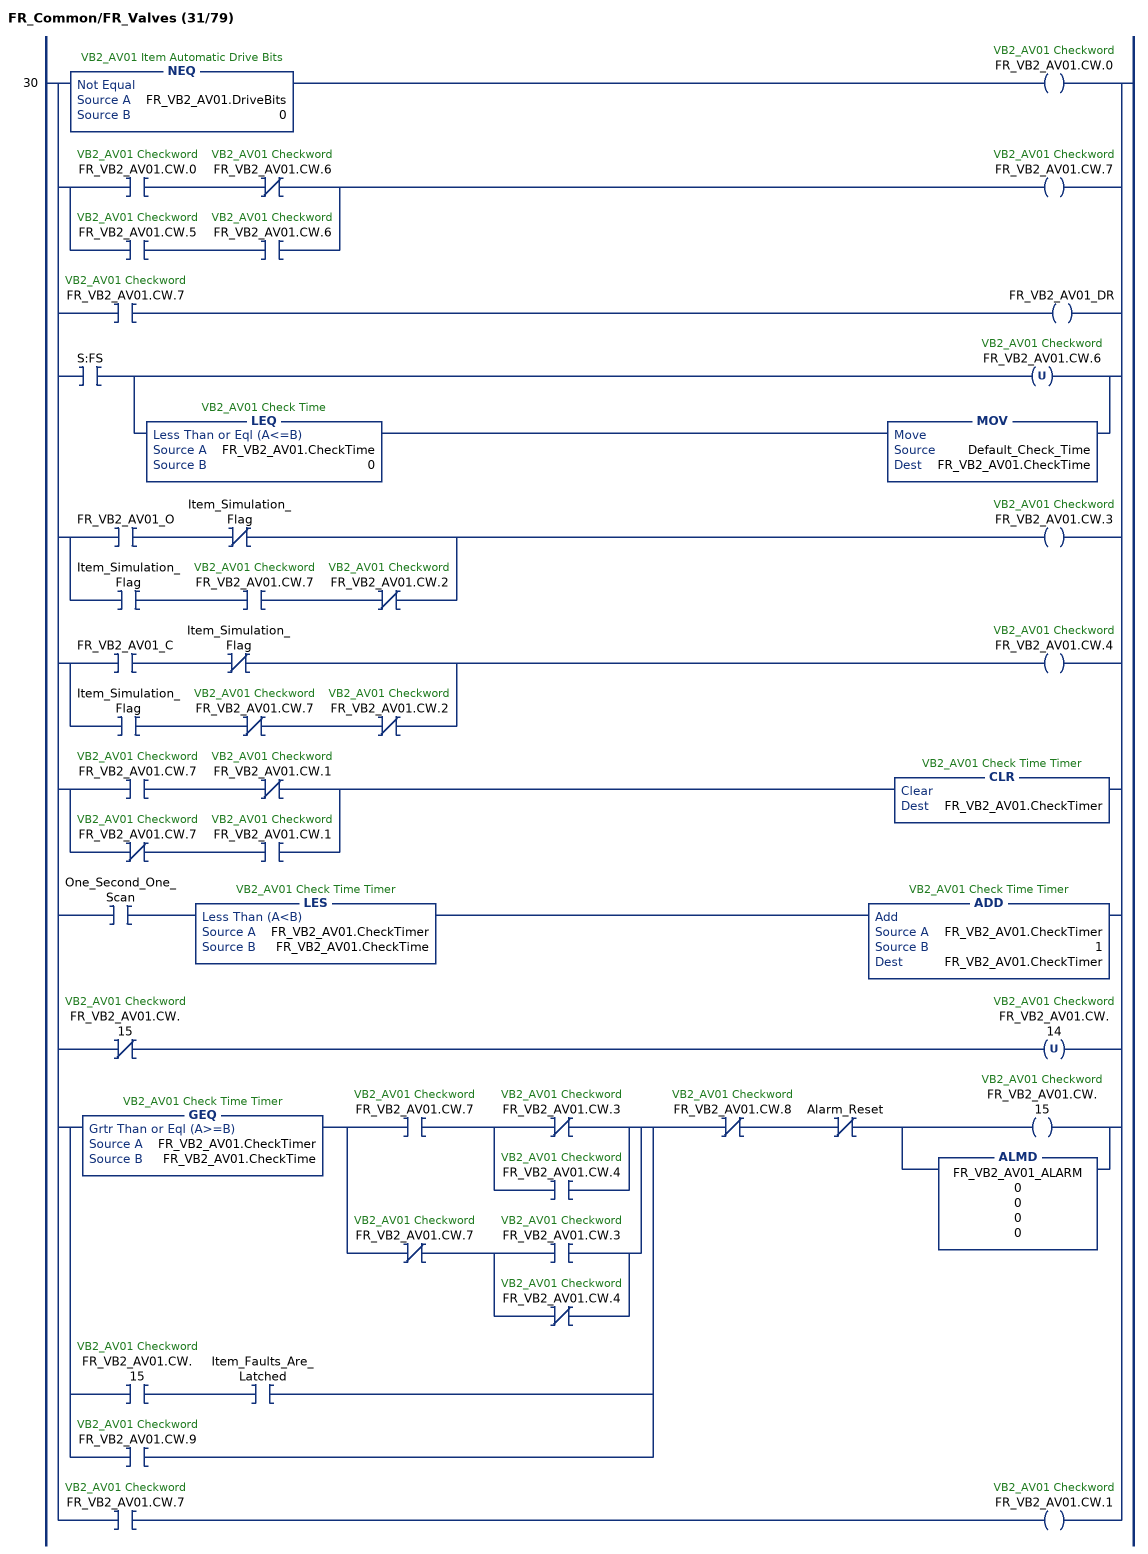
   30: [NEQ(FR_VB2_AV01.DriveBits,0) OTE(FR_VB2_AV01.CW.0) ,[XIC(FR_VB2_AV01.CW.0) XIO(FR_VB2_AV01.CW.6) ,XIC(FR_VB2_AV01.CW.5) XIC(FR_VB2_AV01.CW.6) ] OTE(FR_VB2_AV01.CW.7) ,XIC(FR_VB2_AV01.CW.7) OTE(FR_VB2_AV01_DR) ,XIC(S:FS) [OTU(FR_VB2_AV01.CW.6) ,LEQ(FR_VB2_AV01.CheckTime,0) MOV(Default_Check_Time,FR_VB2_AV01.CheckTime) ] ,[[XIC(FR_VB2_AV01_O) XIO(Item_Simulation_Flag) ,XIC(Item_Simulation_Flag) XIC(FR_VB2_AV01.CW.7) XIO(FR_VB2_AV01.CW.2) ] OTE(FR_VB2_AV01.CW.3) ,[XIC(FR_VB2_AV01_C) XIO(Item_Simulation_Flag) ,XIC(Item_Simulation_Flag) XIO(FR_VB2_AV01.CW.7) XIO(FR_VB2_AV01.CW.2) ] OTE(FR_VB2_AV01.CW.4) ] ,[XIC(FR_VB2_AV01.CW.7) XIO(FR_VB2_AV01.CW.1) ,XIO(FR_VB2_AV01.CW.7) XIC(FR_VB2_AV01.CW.1) ] CLR(FR_VB2_AV01.CheckTimer) ,XIC(One_Second_One_Scan) LES(FR_VB2_AV01.CheckTimer,FR_VB2_AV01.CheckTime) ADD(FR_VB2_AV01.CheckTimer,1,FR_VB2_AV01.CheckTimer) ,XIO(FR_VB2_AV01.CW.15) OTU(FR_VB2_AV01.CW.14) ,[GEQ(FR_VB2_AV01.CheckTimer,FR_VB2_AV01.CheckTime) [XIC(FR_VB2_AV01.CW.7) [XIO(FR_VB2_AV01.CW.3) ,XIC(FR_VB2_AV01.CW.4) ] ,XIO(FR_VB2_AV01.CW.7) [XIC(FR_VB2_AV01.CW.3) ,XIO(FR_VB2_AV01.CW.4) ] ] ,XIC(FR_VB2_AV01.CW.15) XIC(Item_Faults_Are_Latched) ,XIC(FR_VB2_AV01.CW.9) ] XIO(FR_VB2_AV01.CW.8) XIO(Alarm_Reset) [OTE(FR_VB2_AV01.CW.15) ,ALMD(FR_VB2_AV01_ALARM,0,0,0,0) ] ,XIC(FR_VB2_AV01.CW.7) OTE(FR_VB2_AV01.CW.1) ];
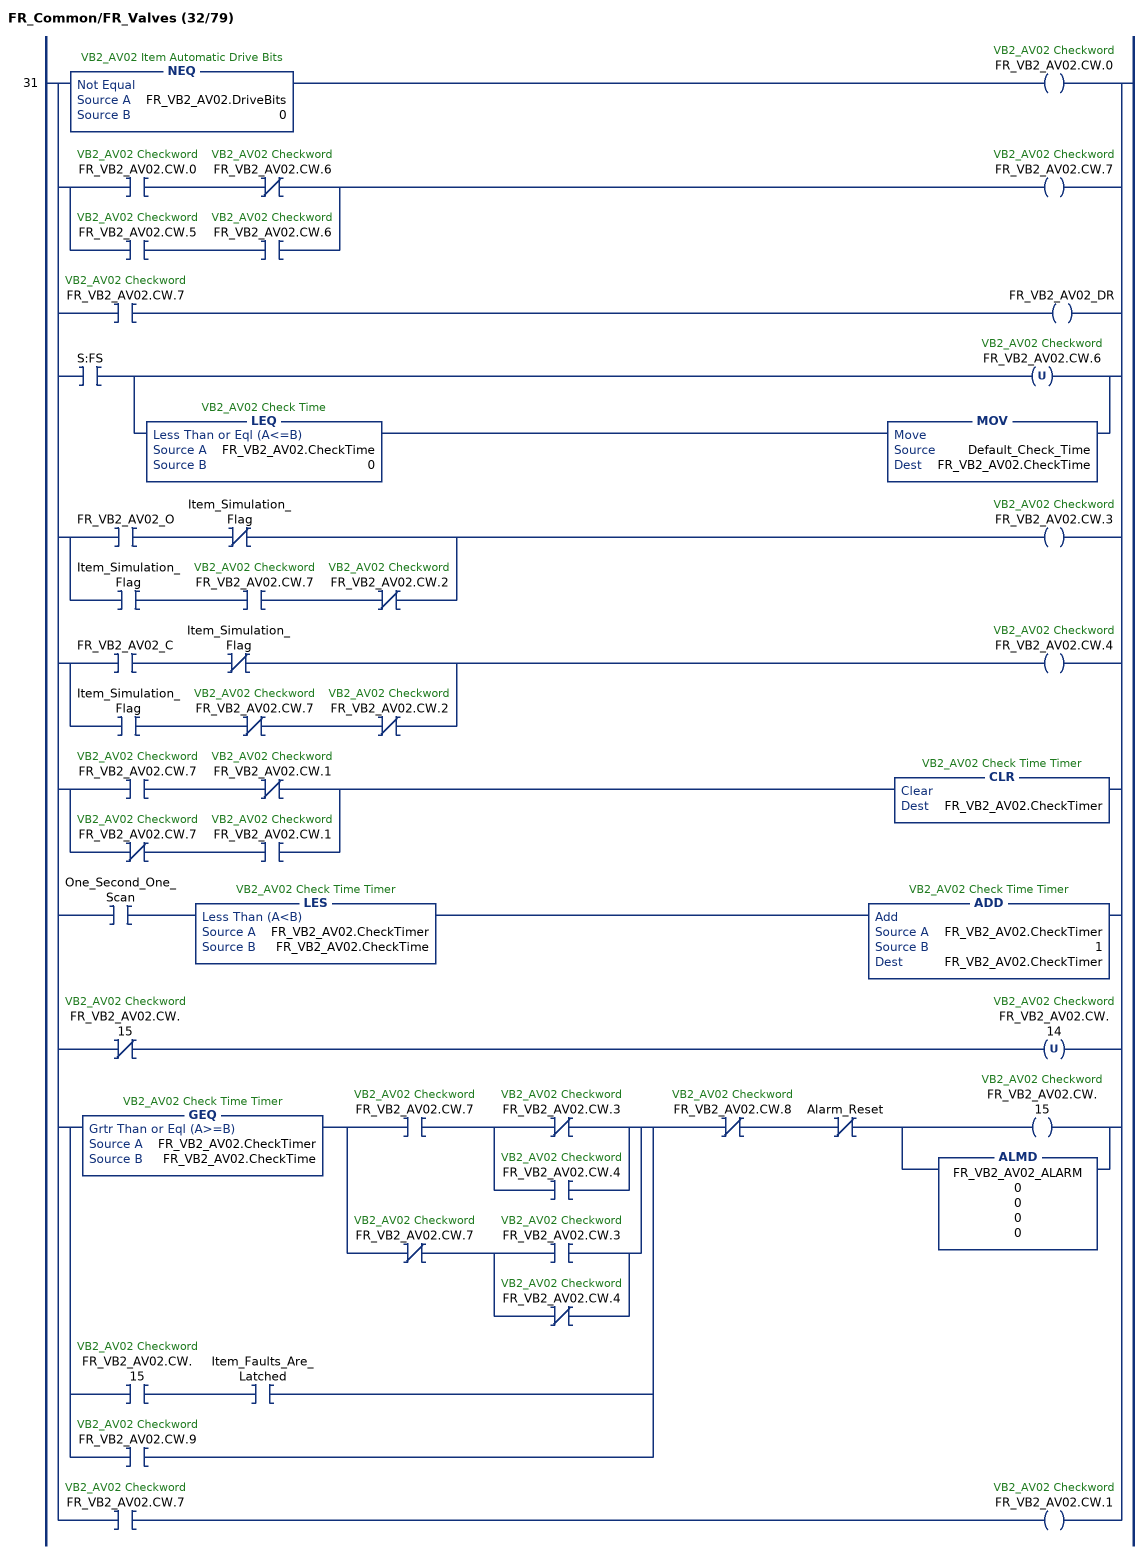
   31: [NEQ(FR_VB2_AV02.DriveBits,0) OTE(FR_VB2_AV02.CW.0) ,[XIC(FR_VB2_AV02.CW.0) XIO(FR_VB2_AV02.CW.6) ,XIC(FR_VB2_AV02.CW.5) XIC(FR_VB2_AV02.CW.6) ] OTE(FR_VB2_AV02.CW.7) ,XIC(FR_VB2_AV02.CW.7) OTE(FR_VB2_AV02_DR) ,XIC(S:FS) [OTU(FR_VB2_AV02.CW.6) ,LEQ(FR_VB2_AV02.CheckTime,0) MOV(Default_Check_Time,FR_VB2_AV02.CheckTime) ] ,[[XIC(FR_VB2_AV02_O) XIO(Item_Simulation_Flag) ,XIC(Item_Simulation_Flag) XIC(FR_VB2_AV02.CW.7) XIO(FR_VB2_AV02.CW.2) ] OTE(FR_VB2_AV02.CW.3) ,[XIC(FR_VB2_AV02_C) XIO(Item_Simulation_Flag) ,XIC(Item_Simulation_Flag) XIO(FR_VB2_AV02.CW.7) XIO(FR_VB2_AV02.CW.2) ] OTE(FR_VB2_AV02.CW.4) ] ,[XIC(FR_VB2_AV02.CW.7) XIO(FR_VB2_AV02.CW.1) ,XIO(FR_VB2_AV02.CW.7) XIC(FR_VB2_AV02.CW.1) ] CLR(FR_VB2_AV02.CheckTimer) ,XIC(One_Second_One_Scan) LES(FR_VB2_AV02.CheckTimer,FR_VB2_AV02.CheckTime) ADD(FR_VB2_AV02.CheckTimer,1,FR_VB2_AV02.CheckTimer) ,XIO(FR_VB2_AV02.CW.15) OTU(FR_VB2_AV02.CW.14) ,[GEQ(FR_VB2_AV02.CheckTimer,FR_VB2_AV02.CheckTime) [XIC(FR_VB2_AV02.CW.7) [XIO(FR_VB2_AV02.CW.3) ,XIC(FR_VB2_AV02.CW.4) ] ,XIO(FR_VB2_AV02.CW.7) [XIC(FR_VB2_AV02.CW.3) ,XIO(FR_VB2_AV02.CW.4) ] ] ,XIC(FR_VB2_AV02.CW.15) XIC(Item_Faults_Are_Latched) ,XIC(FR_VB2_AV02.CW.9) ] XIO(FR_VB2_AV02.CW.8) XIO(Alarm_Reset) [OTE(FR_VB2_AV02.CW.15) ,ALMD(FR_VB2_AV02_ALARM,0,0,0,0) ] ,XIC(FR_VB2_AV02.CW.7) OTE(FR_VB2_AV02.CW.1) ];
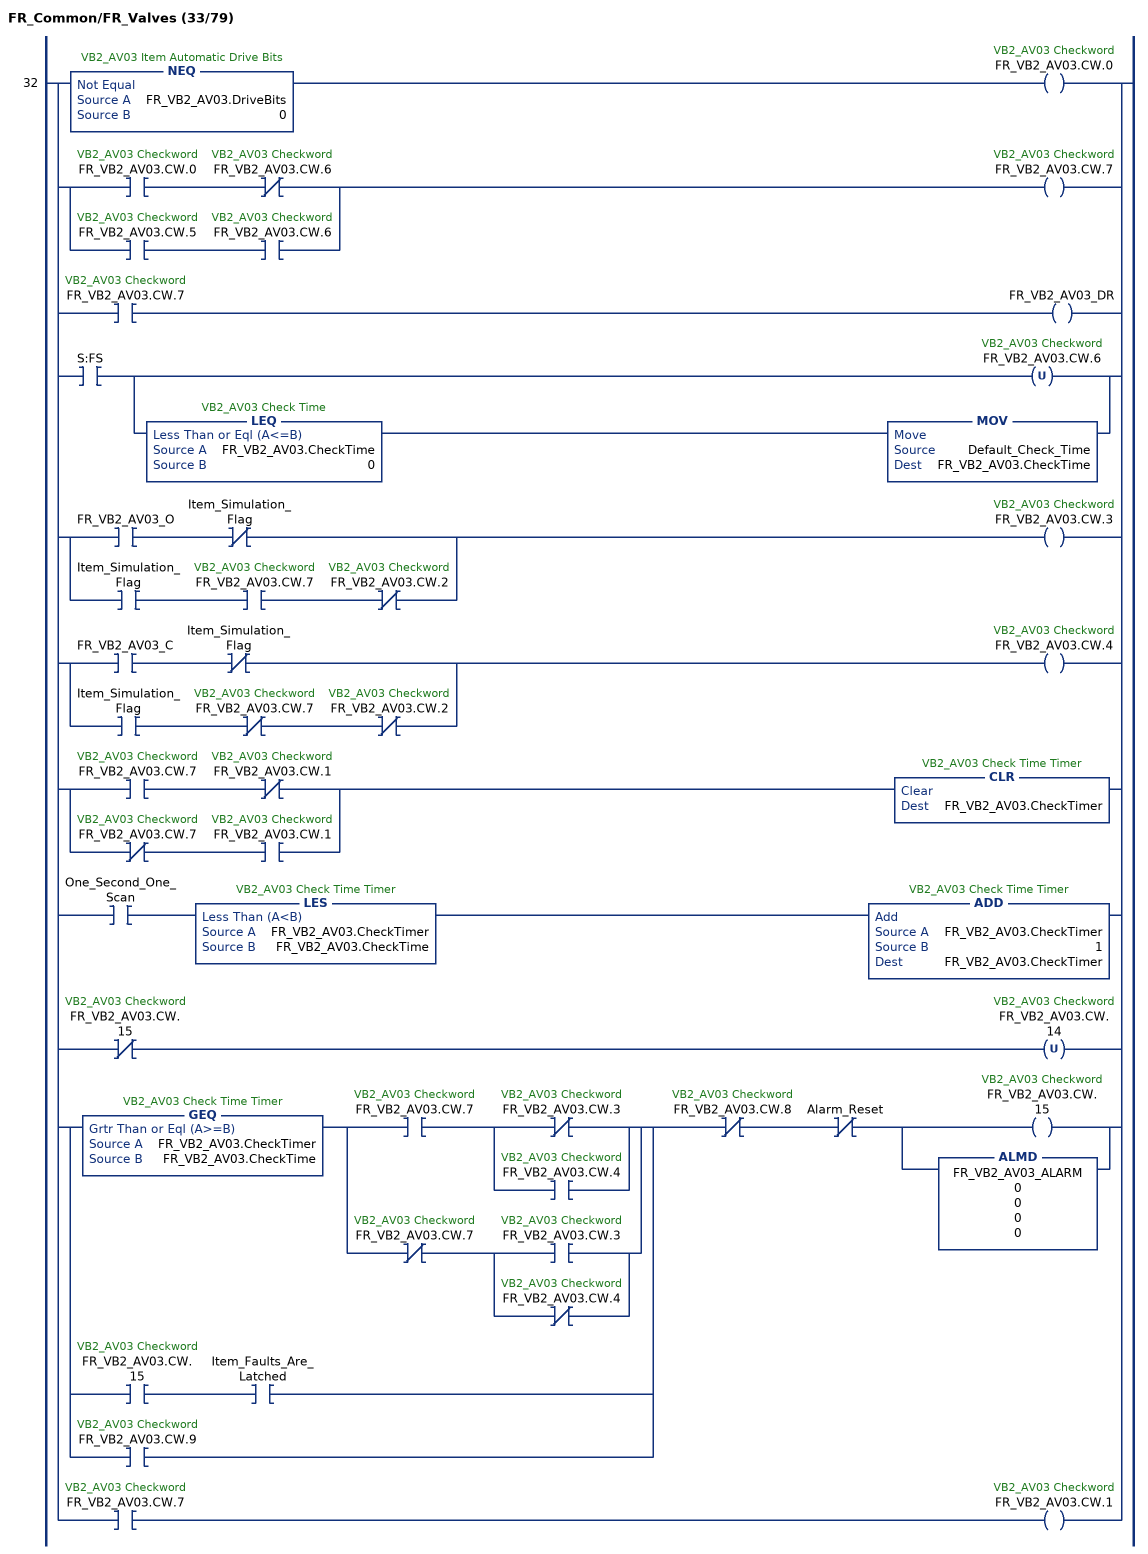
   32: [NEQ(FR_VB2_AV03.DriveBits,0) OTE(FR_VB2_AV03.CW.0) ,[XIC(FR_VB2_AV03.CW.0) XIO(FR_VB2_AV03.CW.6) ,XIC(FR_VB2_AV03.CW.5) XIC(FR_VB2_AV03.CW.6) ] OTE(FR_VB2_AV03.CW.7) ,XIC(FR_VB2_AV03.CW.7) OTE(FR_VB2_AV03_DR) ,XIC(S:FS) [OTU(FR_VB2_AV03.CW.6) ,LEQ(FR_VB2_AV03.CheckTime,0) MOV(Default_Check_Time,FR_VB2_AV03.CheckTime) ] ,[[XIC(FR_VB2_AV03_O) XIO(Item_Simulation_Flag) ,XIC(Item_Simulation_Flag) XIC(FR_VB2_AV03.CW.7) XIO(FR_VB2_AV03.CW.2) ] OTE(FR_VB2_AV03.CW.3) ,[XIC(FR_VB2_AV03_C) XIO(Item_Simulation_Flag) ,XIC(Item_Simulation_Flag) XIO(FR_VB2_AV03.CW.7) XIO(FR_VB2_AV03.CW.2) ] OTE(FR_VB2_AV03.CW.4) ] ,[XIC(FR_VB2_AV03.CW.7) XIO(FR_VB2_AV03.CW.1) ,XIO(FR_VB2_AV03.CW.7) XIC(FR_VB2_AV03.CW.1) ] CLR(FR_VB2_AV03.CheckTimer) ,XIC(One_Second_One_Scan) LES(FR_VB2_AV03.CheckTimer,FR_VB2_AV03.CheckTime) ADD(FR_VB2_AV03.CheckTimer,1,FR_VB2_AV03.CheckTimer) ,XIO(FR_VB2_AV03.CW.15) OTU(FR_VB2_AV03.CW.14) ,[GEQ(FR_VB2_AV03.CheckTimer,FR_VB2_AV03.CheckTime) [XIC(FR_VB2_AV03.CW.7) [XIO(FR_VB2_AV03.CW.3) ,XIC(FR_VB2_AV03.CW.4) ] ,XIO(FR_VB2_AV03.CW.7) [XIC(FR_VB2_AV03.CW.3) ,XIO(FR_VB2_AV03.CW.4) ] ] ,XIC(FR_VB2_AV03.CW.15) XIC(Item_Faults_Are_Latched) ,XIC(FR_VB2_AV03.CW.9) ] XIO(FR_VB2_AV03.CW.8) XIO(Alarm_Reset) [OTE(FR_VB2_AV03.CW.15) ,ALMD(FR_VB2_AV03_ALARM,0,0,0,0) ] ,XIC(FR_VB2_AV03.CW.7) OTE(FR_VB2_AV03.CW.1) ];
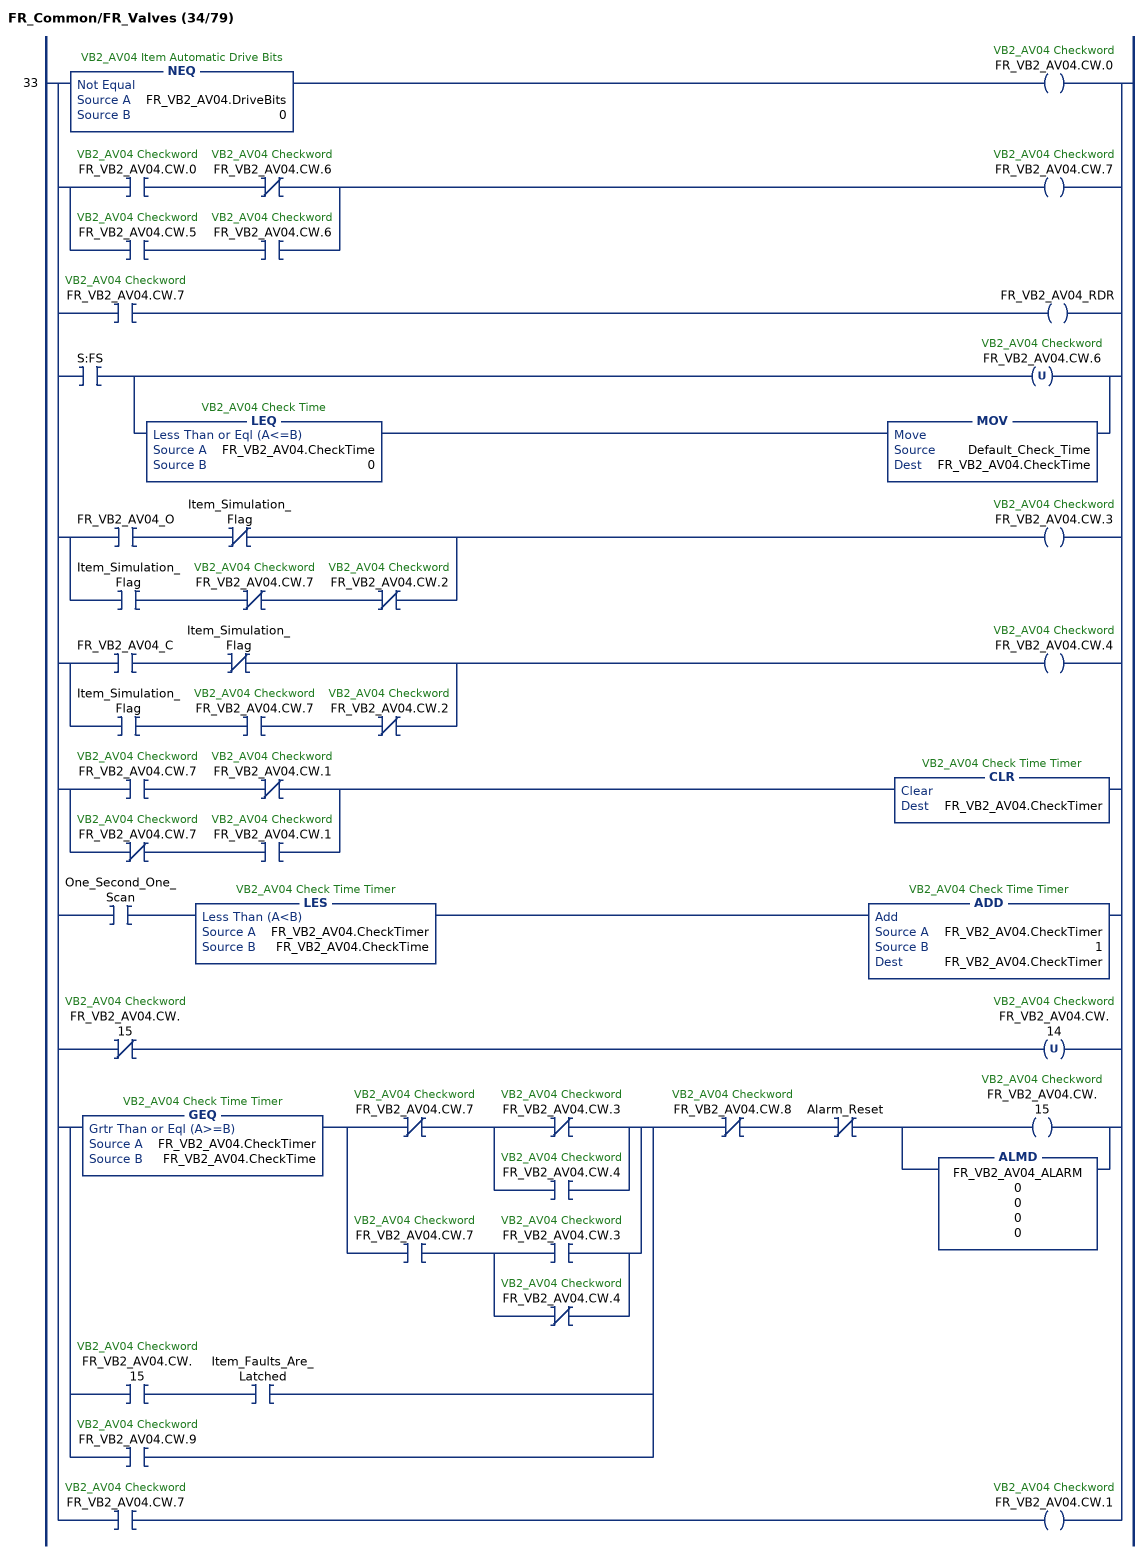
   33: [NEQ(FR_VB2_AV04.DriveBits,0) OTE(FR_VB2_AV04.CW.0) ,[XIC(FR_VB2_AV04.CW.0) XIO(FR_VB2_AV04.CW.6) ,XIC(FR_VB2_AV04.CW.5) XIC(FR_VB2_AV04.CW.6) ] OTE(FR_VB2_AV04.CW.7) ,XIC(FR_VB2_AV04.CW.7) OTE(FR_VB2_AV04_RDR) ,XIC(S:FS) [OTU(FR_VB2_AV04.CW.6) ,LEQ(FR_VB2_AV04.CheckTime,0) MOV(Default_Check_Time,FR_VB2_AV04.CheckTime) ] ,[[XIC(FR_VB2_AV04_O) XIO(Item_Simulation_Flag) ,XIC(Item_Simulation_Flag) XIO(FR_VB2_AV04.CW.7) XIO(FR_VB2_AV04.CW.2) ] OTE(FR_VB2_AV04.CW.3) ,[XIC(FR_VB2_AV04_C) XIO(Item_Simulation_Flag) ,XIC(Item_Simulation_Flag) XIC(FR_VB2_AV04.CW.7) XIO(FR_VB2_AV04.CW.2) ] OTE(FR_VB2_AV04.CW.4) ] ,[XIC(FR_VB2_AV04.CW.7) XIO(FR_VB2_AV04.CW.1) ,XIO(FR_VB2_AV04.CW.7) XIC(FR_VB2_AV04.CW.1) ] CLR(FR_VB2_AV04.CheckTimer) ,XIC(One_Second_One_Scan) LES(FR_VB2_AV04.CheckTimer,FR_VB2_AV04.CheckTime) ADD(FR_VB2_AV04.CheckTimer,1,FR_VB2_AV04.CheckTimer) ,XIO(FR_VB2_AV04.CW.15) OTU(FR_VB2_AV04.CW.14) ,[GEQ(FR_VB2_AV04.CheckTimer,FR_VB2_AV04.CheckTime) [XIO(FR_VB2_AV04.CW.7) [XIO(FR_VB2_AV04.CW.3) ,XIC(FR_VB2_AV04.CW.4) ] ,XIC(FR_VB2_AV04.CW.7) [XIC(FR_VB2_AV04.CW.3) ,XIO(FR_VB2_AV04.CW.4) ] ] ,XIC(FR_VB2_AV04.CW.15) XIC(Item_Faults_Are_Latched) ,XIC(FR_VB2_AV04.CW.9) ] XIO(FR_VB2_AV04.CW.8) XIO(Alarm_Reset) [OTE(FR_VB2_AV04.CW.15) ,ALMD(FR_VB2_AV04_ALARM,0,0,0,0) ] ,XIC(FR_VB2_AV04.CW.7) OTE(FR_VB2_AV04.CW.1) ];
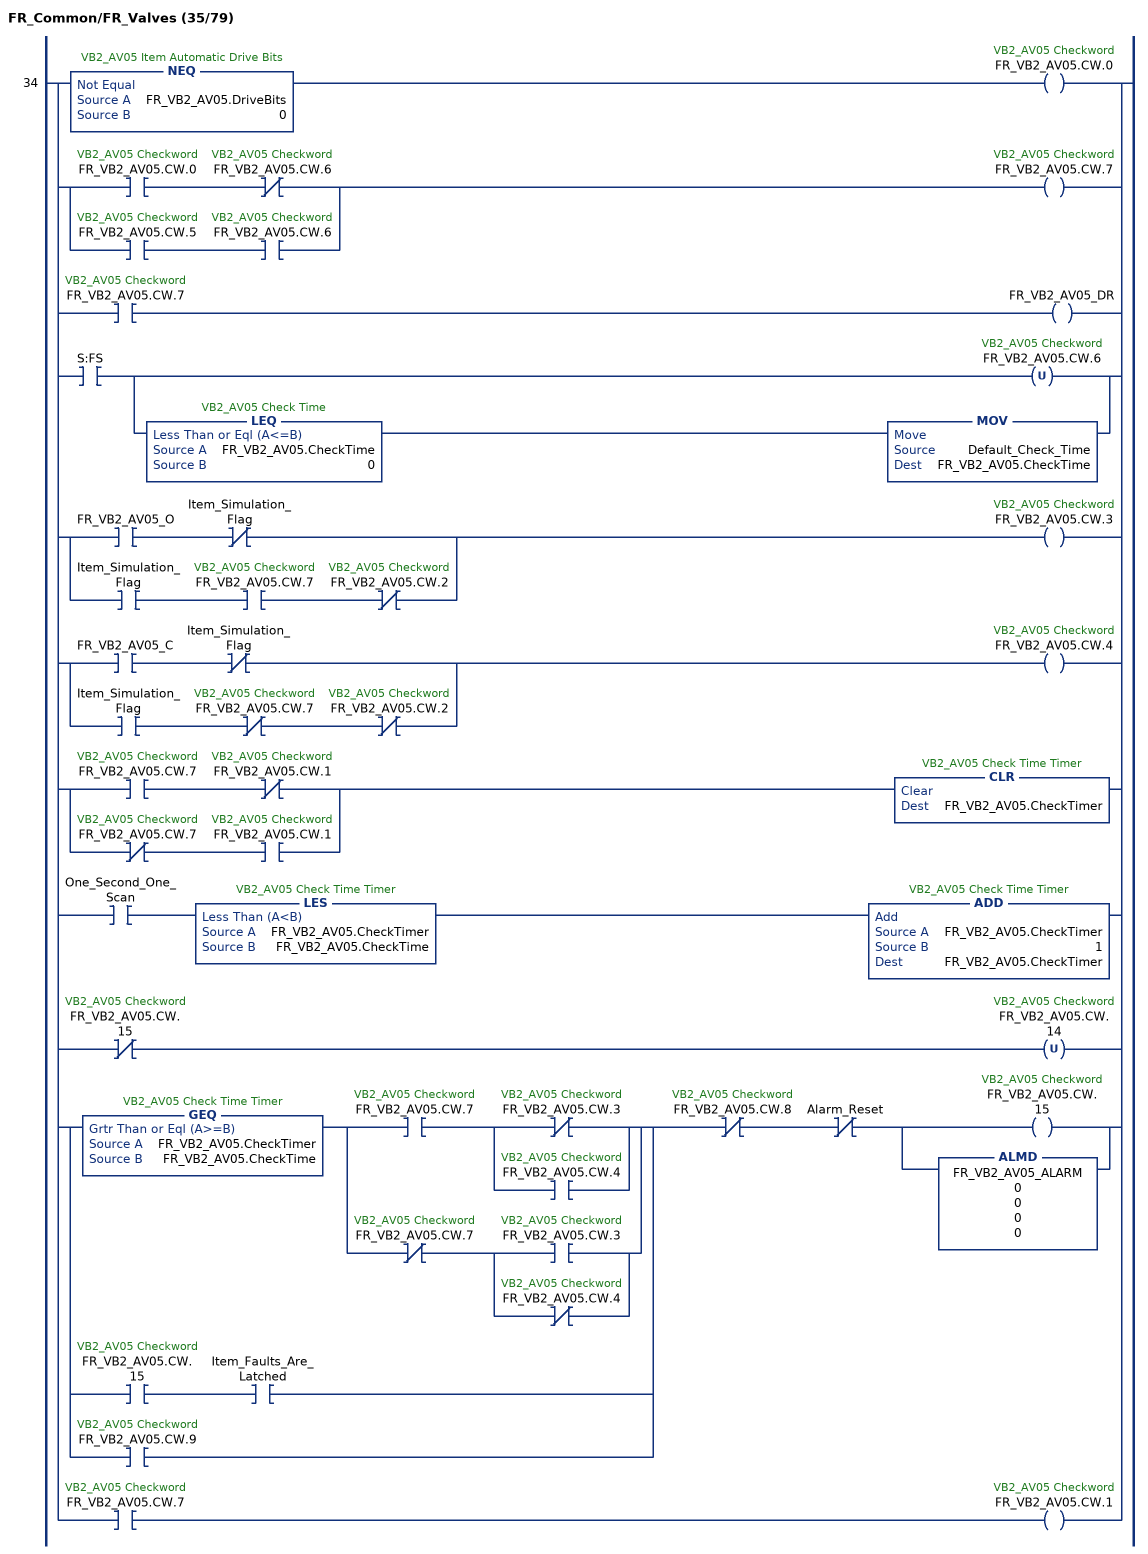
   34: [NEQ(FR_VB2_AV05.DriveBits,0) OTE(FR_VB2_AV05.CW.0) ,[XIC(FR_VB2_AV05.CW.0) XIO(FR_VB2_AV05.CW.6) ,XIC(FR_VB2_AV05.CW.5) XIC(FR_VB2_AV05.CW.6) ] OTE(FR_VB2_AV05.CW.7) ,XIC(FR_VB2_AV05.CW.7) OTE(FR_VB2_AV05_DR) ,XIC(S:FS) [OTU(FR_VB2_AV05.CW.6) ,LEQ(FR_VB2_AV05.CheckTime,0) MOV(Default_Check_Time,FR_VB2_AV05.CheckTime) ] ,[[XIC(FR_VB2_AV05_O) XIO(Item_Simulation_Flag) ,XIC(Item_Simulation_Flag) XIC(FR_VB2_AV05.CW.7) XIO(FR_VB2_AV05.CW.2) ] OTE(FR_VB2_AV05.CW.3) ,[XIC(FR_VB2_AV05_C) XIO(Item_Simulation_Flag) ,XIC(Item_Simulation_Flag) XIO(FR_VB2_AV05.CW.7) XIO(FR_VB2_AV05.CW.2) ] OTE(FR_VB2_AV05.CW.4) ] ,[XIC(FR_VB2_AV05.CW.7) XIO(FR_VB2_AV05.CW.1) ,XIO(FR_VB2_AV05.CW.7) XIC(FR_VB2_AV05.CW.1) ] CLR(FR_VB2_AV05.CheckTimer) ,XIC(One_Second_One_Scan) LES(FR_VB2_AV05.CheckTimer,FR_VB2_AV05.CheckTime) ADD(FR_VB2_AV05.CheckTimer,1,FR_VB2_AV05.CheckTimer) ,XIO(FR_VB2_AV05.CW.15) OTU(FR_VB2_AV05.CW.14) ,[GEQ(FR_VB2_AV05.CheckTimer,FR_VB2_AV05.CheckTime) [XIC(FR_VB2_AV05.CW.7) [XIO(FR_VB2_AV05.CW.3) ,XIC(FR_VB2_AV05.CW.4) ] ,XIO(FR_VB2_AV05.CW.7) [XIC(FR_VB2_AV05.CW.3) ,XIO(FR_VB2_AV05.CW.4) ] ] ,XIC(FR_VB2_AV05.CW.15) XIC(Item_Faults_Are_Latched) ,XIC(FR_VB2_AV05.CW.9) ] XIO(FR_VB2_AV05.CW.8) XIO(Alarm_Reset) [OTE(FR_VB2_AV05.CW.15) ,ALMD(FR_VB2_AV05_ALARM,0,0,0,0) ] ,XIC(FR_VB2_AV05.CW.7) OTE(FR_VB2_AV05.CW.1) ];
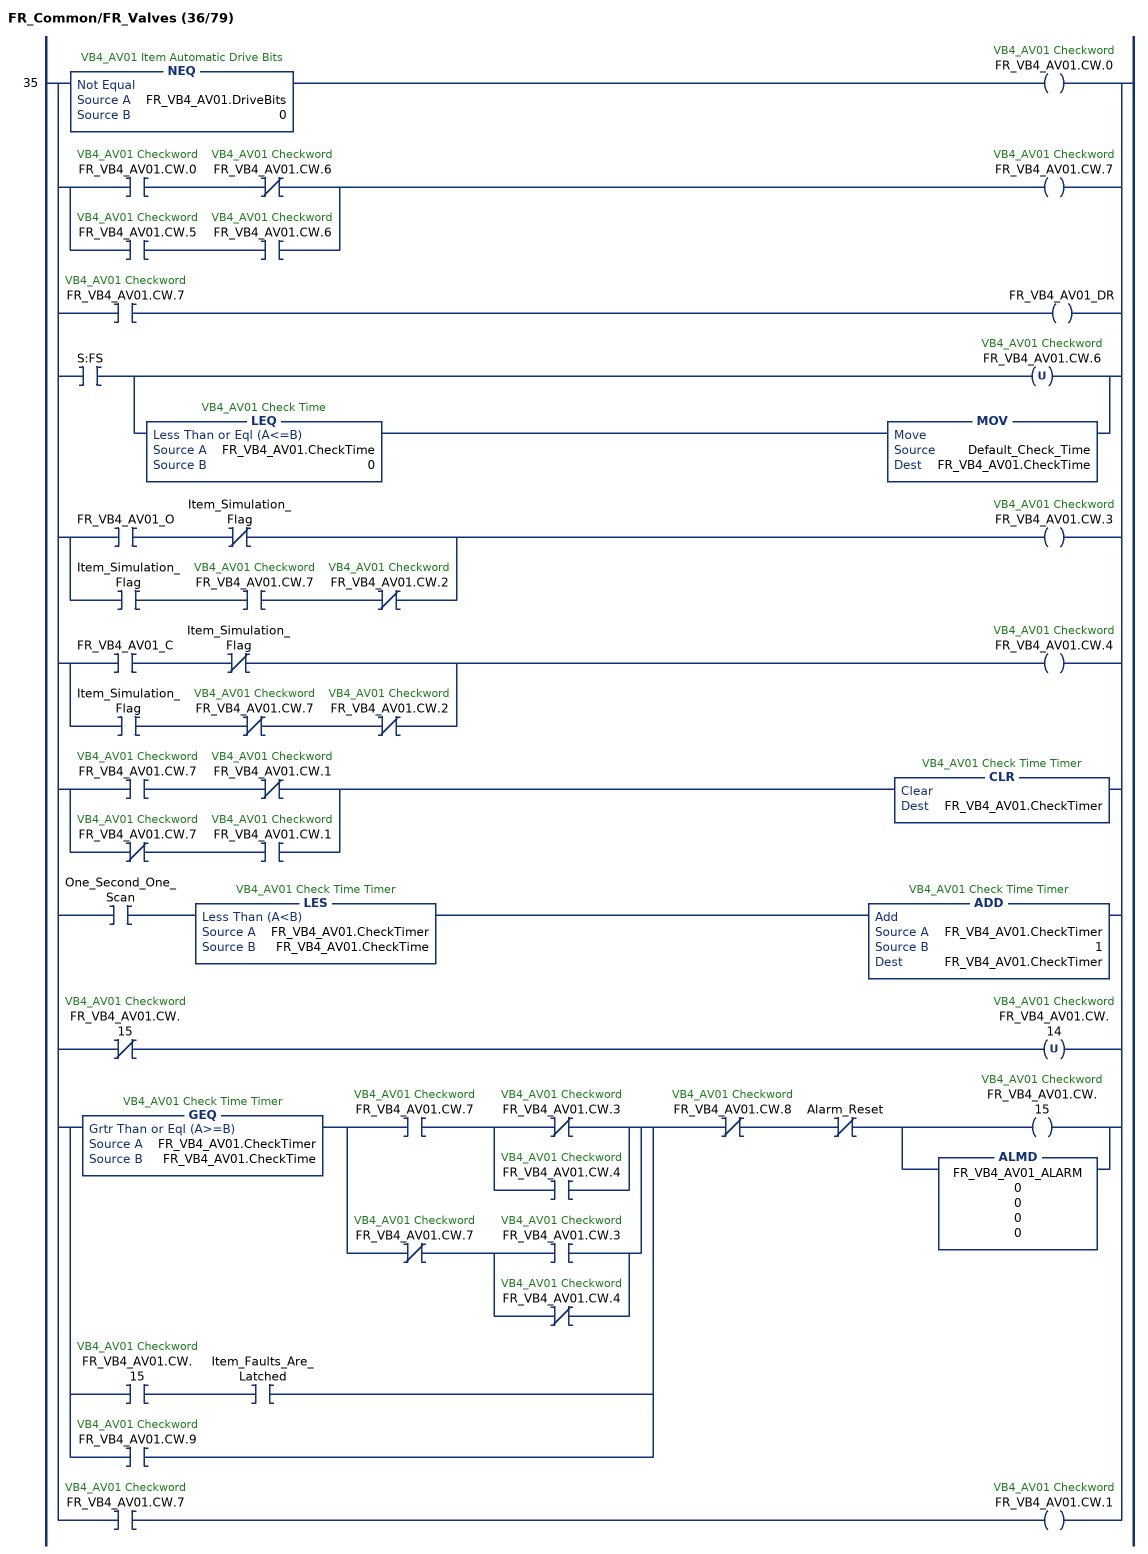
   35: [NEQ(FR_VB4_AV01.DriveBits,0) OTE(FR_VB4_AV01.CW.0) ,[XIC(FR_VB4_AV01.CW.0) XIO(FR_VB4_AV01.CW.6) ,XIC(FR_VB4_AV01.CW.5) XIC(FR_VB4_AV01.CW.6) ] OTE(FR_VB4_AV01.CW.7) ,XIC(FR_VB4_AV01.CW.7) OTE(FR_VB4_AV01_DR) ,XIC(S:FS) [OTU(FR_VB4_AV01.CW.6) ,LEQ(FR_VB4_AV01.CheckTime,0) MOV(Default_Check_Time,FR_VB4_AV01.CheckTime) ] ,[[XIC(FR_VB4_AV01_O) XIO(Item_Simulation_Flag) ,XIC(Item_Simulation_Flag) XIC(FR_VB4_AV01.CW.7) XIO(FR_VB4_AV01.CW.2) ] OTE(FR_VB4_AV01.CW.3) ,[XIC(FR_VB4_AV01_C) XIO(Item_Simulation_Flag) ,XIC(Item_Simulation_Flag) XIO(FR_VB4_AV01.CW.7) XIO(FR_VB4_AV01.CW.2) ] OTE(FR_VB4_AV01.CW.4) ] ,[XIC(FR_VB4_AV01.CW.7) XIO(FR_VB4_AV01.CW.1) ,XIO(FR_VB4_AV01.CW.7) XIC(FR_VB4_AV01.CW.1) ] CLR(FR_VB4_AV01.CheckTimer) ,XIC(One_Second_One_Scan) LES(FR_VB4_AV01.CheckTimer,FR_VB4_AV01.CheckTime) ADD(FR_VB4_AV01.CheckTimer,1,FR_VB4_AV01.CheckTimer) ,XIO(FR_VB4_AV01.CW.15) OTU(FR_VB4_AV01.CW.14) ,[GEQ(FR_VB4_AV01.CheckTimer,FR_VB4_AV01.CheckTime) [XIC(FR_VB4_AV01.CW.7) [XIO(FR_VB4_AV01.CW.3) ,XIC(FR_VB4_AV01.CW.4) ] ,XIO(FR_VB4_AV01.CW.7) [XIC(FR_VB4_AV01.CW.3) ,XIO(FR_VB4_AV01.CW.4) ] ] ,XIC(FR_VB4_AV01.CW.15) XIC(Item_Faults_Are_Latched) ,XIC(FR_VB4_AV01.CW.9) ] XIO(FR_VB4_AV01.CW.8) XIO(Alarm_Reset) [OTE(FR_VB4_AV01.CW.15) ,ALMD(FR_VB4_AV01_ALARM,0,0,0,0) ] ,XIC(FR_VB4_AV01.CW.7) OTE(FR_VB4_AV01.CW.1) ];
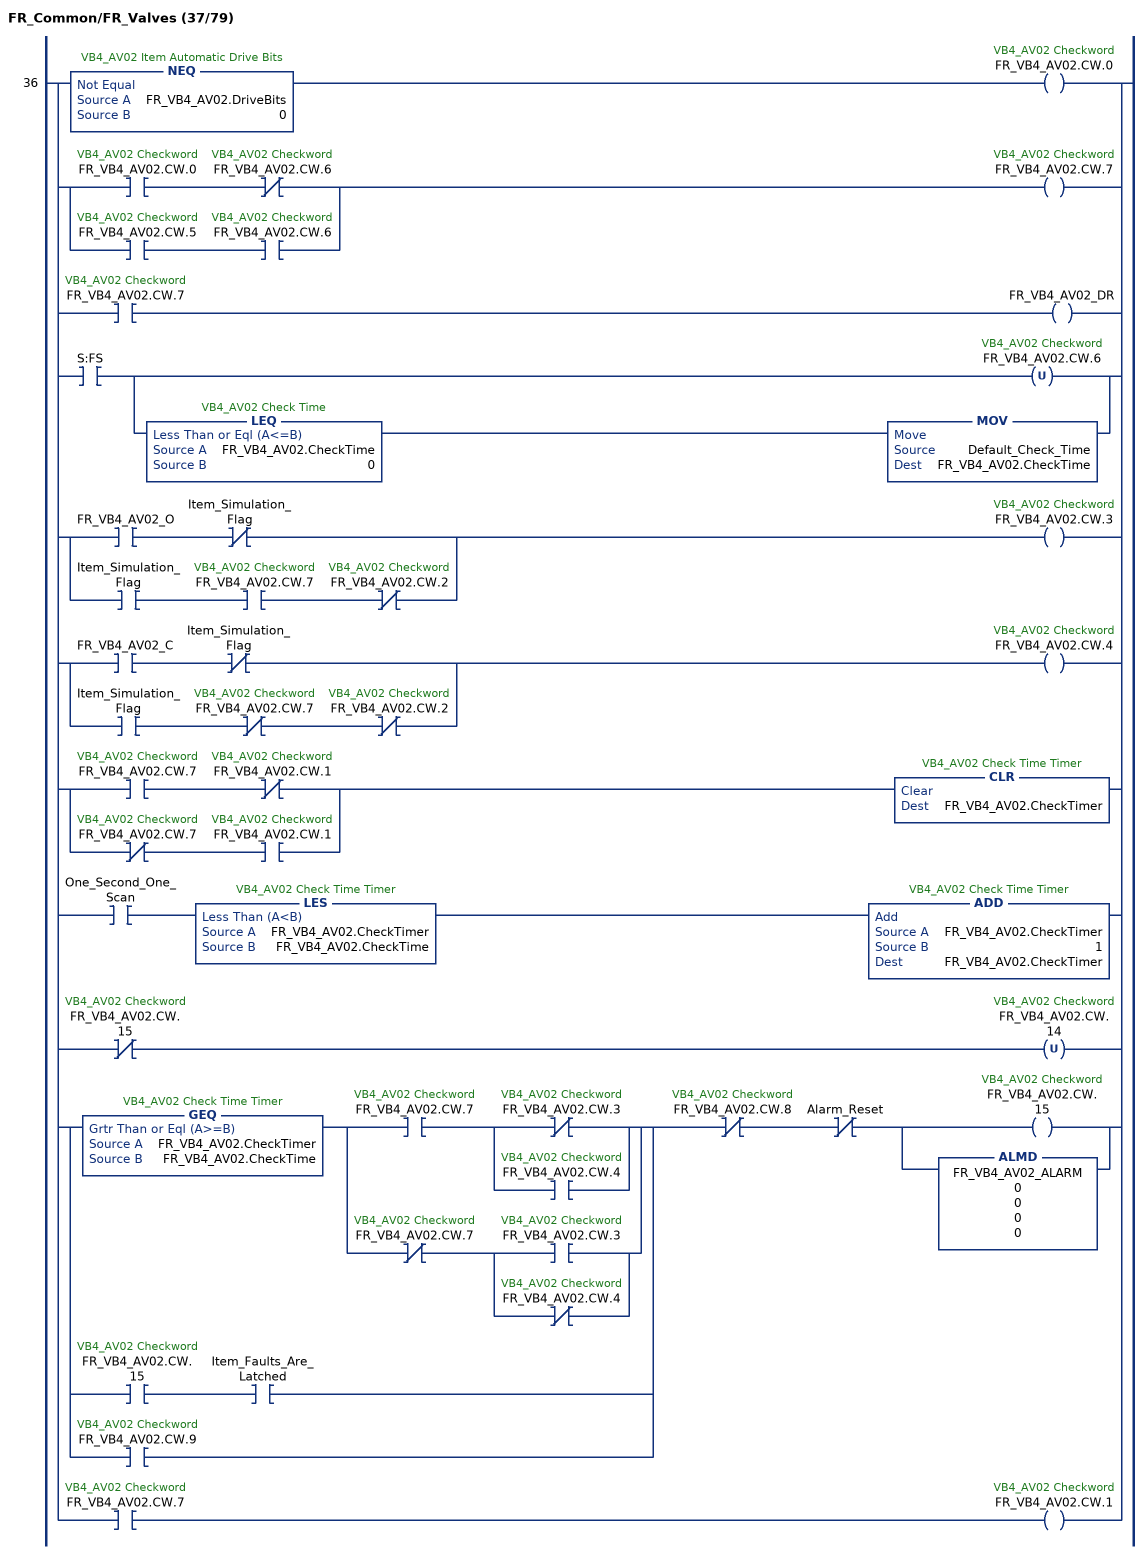
   36: [NEQ(FR_VB4_AV02.DriveBits,0) OTE(FR_VB4_AV02.CW.0) ,[XIC(FR_VB4_AV02.CW.0) XIO(FR_VB4_AV02.CW.6) ,XIC(FR_VB4_AV02.CW.5) XIC(FR_VB4_AV02.CW.6) ] OTE(FR_VB4_AV02.CW.7) ,XIC(FR_VB4_AV02.CW.7) OTE(FR_VB4_AV02_DR) ,XIC(S:FS) [OTU(FR_VB4_AV02.CW.6) ,LEQ(FR_VB4_AV02.CheckTime,0) MOV(Default_Check_Time,FR_VB4_AV02.CheckTime) ] ,[[XIC(FR_VB4_AV02_O) XIO(Item_Simulation_Flag) ,XIC(Item_Simulation_Flag) XIC(FR_VB4_AV02.CW.7) XIO(FR_VB4_AV02.CW.2) ] OTE(FR_VB4_AV02.CW.3) ,[XIC(FR_VB4_AV02_C) XIO(Item_Simulation_Flag) ,XIC(Item_Simulation_Flag) XIO(FR_VB4_AV02.CW.7) XIO(FR_VB4_AV02.CW.2) ] OTE(FR_VB4_AV02.CW.4) ] ,[XIC(FR_VB4_AV02.CW.7) XIO(FR_VB4_AV02.CW.1) ,XIO(FR_VB4_AV02.CW.7) XIC(FR_VB4_AV02.CW.1) ] CLR(FR_VB4_AV02.CheckTimer) ,XIC(One_Second_One_Scan) LES(FR_VB4_AV02.CheckTimer,FR_VB4_AV02.CheckTime) ADD(FR_VB4_AV02.CheckTimer,1,FR_VB4_AV02.CheckTimer) ,XIO(FR_VB4_AV02.CW.15) OTU(FR_VB4_AV02.CW.14) ,[GEQ(FR_VB4_AV02.CheckTimer,FR_VB4_AV02.CheckTime) [XIC(FR_VB4_AV02.CW.7) [XIO(FR_VB4_AV02.CW.3) ,XIC(FR_VB4_AV02.CW.4) ] ,XIO(FR_VB4_AV02.CW.7) [XIC(FR_VB4_AV02.CW.3) ,XIO(FR_VB4_AV02.CW.4) ] ] ,XIC(FR_VB4_AV02.CW.15) XIC(Item_Faults_Are_Latched) ,XIC(FR_VB4_AV02.CW.9) ] XIO(FR_VB4_AV02.CW.8) XIO(Alarm_Reset) [OTE(FR_VB4_AV02.CW.15) ,ALMD(FR_VB4_AV02_ALARM,0,0,0,0) ] ,XIC(FR_VB4_AV02.CW.7) OTE(FR_VB4_AV02.CW.1) ];
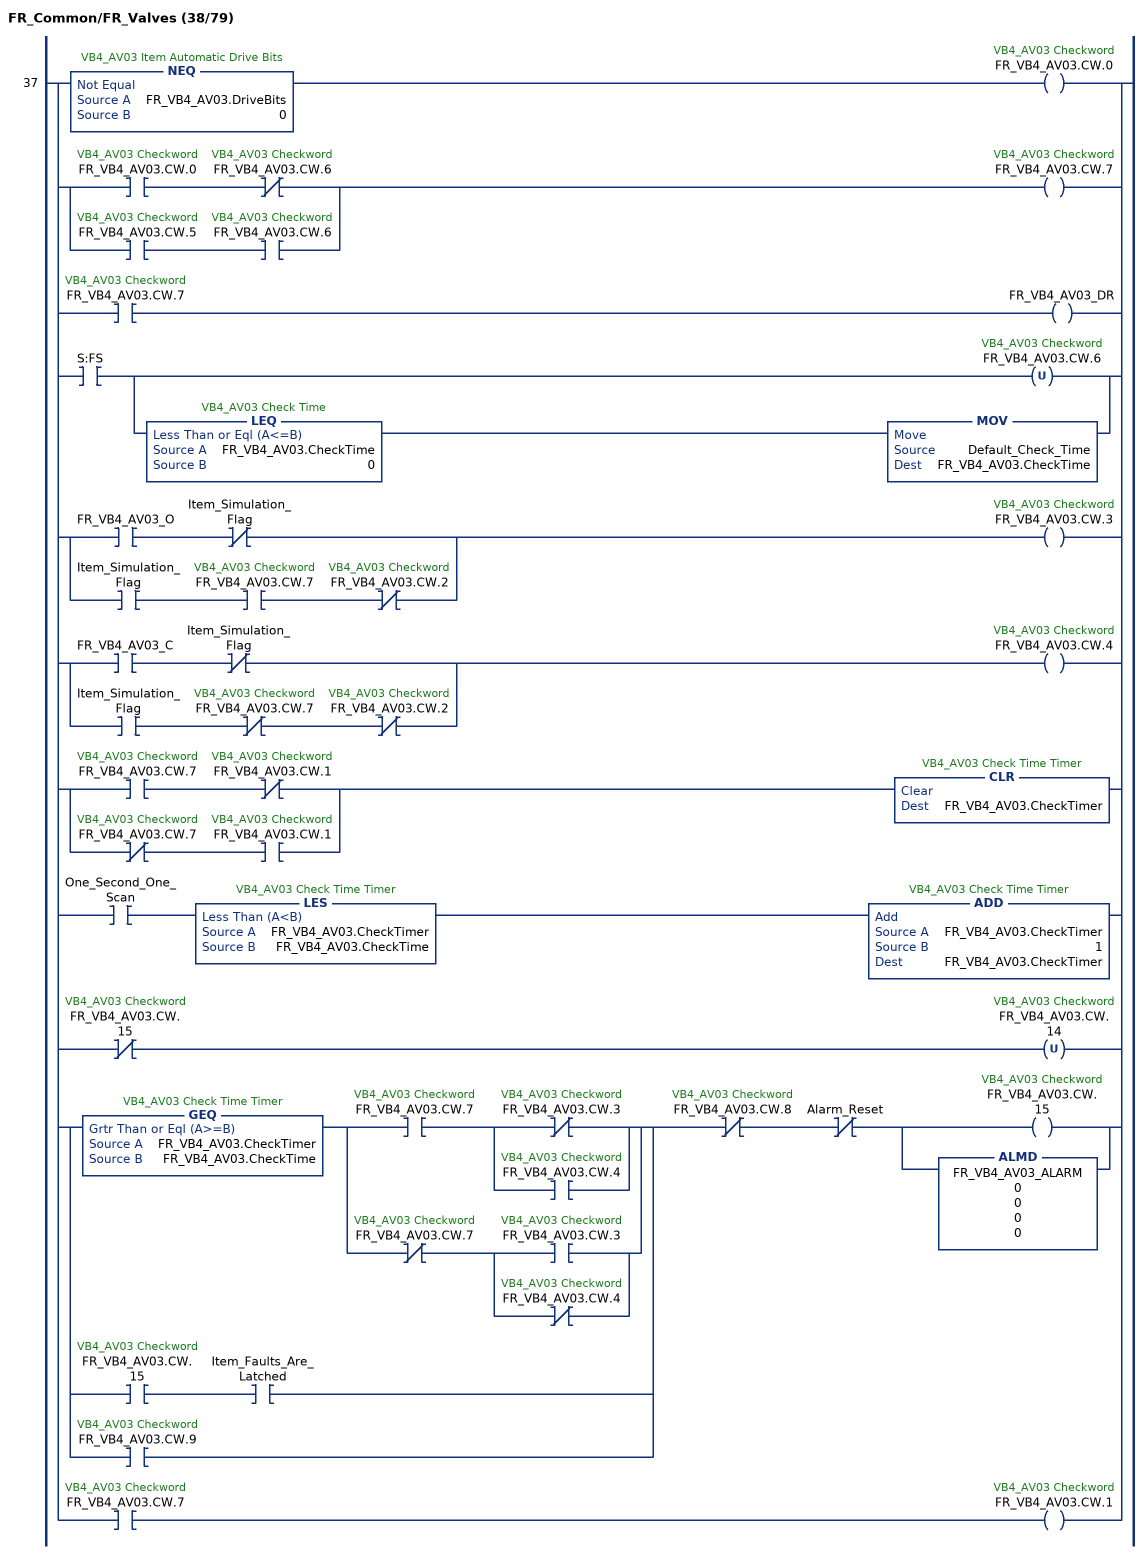
   37: [NEQ(FR_VB4_AV03.DriveBits,0) OTE(FR_VB4_AV03.CW.0) ,[XIC(FR_VB4_AV03.CW.0) XIO(FR_VB4_AV03.CW.6) ,XIC(FR_VB4_AV03.CW.5) XIC(FR_VB4_AV03.CW.6) ] OTE(FR_VB4_AV03.CW.7) ,XIC(FR_VB4_AV03.CW.7) OTE(FR_VB4_AV03_DR) ,XIC(S:FS) [OTU(FR_VB4_AV03.CW.6) ,LEQ(FR_VB4_AV03.CheckTime,0) MOV(Default_Check_Time,FR_VB4_AV03.CheckTime) ] ,[[XIC(FR_VB4_AV03_O) XIO(Item_Simulation_Flag) ,XIC(Item_Simulation_Flag) XIC(FR_VB4_AV03.CW.7) XIO(FR_VB4_AV03.CW.2) ] OTE(FR_VB4_AV03.CW.3) ,[XIC(FR_VB4_AV03_C) XIO(Item_Simulation_Flag) ,XIC(Item_Simulation_Flag) XIO(FR_VB4_AV03.CW.7) XIO(FR_VB4_AV03.CW.2) ] OTE(FR_VB4_AV03.CW.4) ] ,[XIC(FR_VB4_AV03.CW.7) XIO(FR_VB4_AV03.CW.1) ,XIO(FR_VB4_AV03.CW.7) XIC(FR_VB4_AV03.CW.1) ] CLR(FR_VB4_AV03.CheckTimer) ,XIC(One_Second_One_Scan) LES(FR_VB4_AV03.CheckTimer,FR_VB4_AV03.CheckTime) ADD(FR_VB4_AV03.CheckTimer,1,FR_VB4_AV03.CheckTimer) ,XIO(FR_VB4_AV03.CW.15) OTU(FR_VB4_AV03.CW.14) ,[GEQ(FR_VB4_AV03.CheckTimer,FR_VB4_AV03.CheckTime) [XIC(FR_VB4_AV03.CW.7) [XIO(FR_VB4_AV03.CW.3) ,XIC(FR_VB4_AV03.CW.4) ] ,XIO(FR_VB4_AV03.CW.7) [XIC(FR_VB4_AV03.CW.3) ,XIO(FR_VB4_AV03.CW.4) ] ] ,XIC(FR_VB4_AV03.CW.15) XIC(Item_Faults_Are_Latched) ,XIC(FR_VB4_AV03.CW.9) ] XIO(FR_VB4_AV03.CW.8) XIO(Alarm_Reset) [OTE(FR_VB4_AV03.CW.15) ,ALMD(FR_VB4_AV03_ALARM,0,0,0,0) ] ,XIC(FR_VB4_AV03.CW.7) OTE(FR_VB4_AV03.CW.1) ];
